// TIA Portal project "Mel7_new" (V15.1) (continued)
   L_1c_18."Индикатор: Обрыв" := FALSE;
   L_1c_18."Индикатор: В норме" := FALSE;
   L_1c_18."Индикатор: HH активирована" := FALSE;
   L_1c_18."Индикатор: H активирована" := FALSE;
   L_1c_18."Индикатор: L активирована" := FALSE;
   L_1c_18."Индикатор: LL активирована" := FALSE;
   L_1c_18."Уставка: MAX" := 450.0;
   L_1c_18."Уставка: MIN" := 0.0;
   L_1c_18."Уставка: HH" := 80.0;
   L_1c_18."Уставка: H" := 70.0;
   L_1c_18."Уставка: L" := 15.0;
   L_1c_18."Уставка: LL" := 10.0;
   L_1c_18."Уставка: Перелёт" := 20.0;
   L_1c_18."Уставка: Недолёт" := 4.0;
   L_1c_18.PV := 0.0813802;
   L_1c_18.Ток := 4.002893;
   L_1c_18.AnimCode := 0;
   L_1c_18.Error := 16#0000;
   L_1c_18.Bipolar := FALSE;
   L_1c_18.Overshoot_MIN := 27649;
   L_1c_18.Undershoot_MAX := -1;
   L_1c_19."Кнопка: Закрыть фейсплату" := FALSE;
   L_1c_19."Кнопка: Активировать HH" := FALSE;
   L_1c_19."Кнопка: Активировать H" := FALSE;
   L_1c_19."Кнопка: Активировать L" := FALSE;
   L_1c_19."Кнопка: Активировать LL" := FALSE;
   L_1c_19."Кнопка: Ремонт" := FALSE;
   L_1c_19.Видимость := FALSE;
   L_1c_19."Индикатор: Зашкал" := FALSE;
   L_1c_19."Индикатор: Перелёт" := FALSE;
   L_1c_19."Авария: Выход за HH" := FALSE;
   L_1c_19."Предупреждение: Выход за H" := FALSE;
   L_1c_19."Предупреждение: Выход за L" := FALSE;
   L_1c_19."Авария: Выход за LL" := FALSE;
   L_1c_19."Индикатор: Недолет" := FALSE;
   L_1c_19."Индикатор: Обрыв" := FALSE;
   L_1c_19."Индикатор: В норме" := FALSE;
   L_1c_19."Индикатор: HH активирована" := FALSE;
   L_1c_19."Индикатор: H активирована" := FALSE;
   L_1c_19."Индикатор: L активирована" := FALSE;
   L_1c_19."Индикатор: LL активирована" := FALSE;
   L_1c_19."Уставка: MAX" := 100.0;
   L_1c_19."Уставка: MIN" := 0.0;
   L_1c_19."Уставка: HH" := 80.0;
   L_1c_19."Уставка: H" := 70.0;
   L_1c_19."Уставка: L" := 15.0;
   L_1c_19."Уставка: LL" := 10.0;
   L_1c_19."Уставка: Перелёт" := 20.0;
   L_1c_19."Уставка: Недолёт" := 4.0;
   L_1c_19.PV := 0.1157407;
   L_1c_19.Ток := 4.018518;
   L_1c_19.AnimCode := 0;
   L_1c_19.Error := 16#0000;
   L_1c_19.Bipolar := FALSE;
   L_1c_19.Overshoot_MIN := 27649;
   L_1c_19.Undershoot_MAX := -1;
   L_1c_20."Кнопка: Закрыть фейсплату" := FALSE;
   L_1c_20."Кнопка: Активировать H" := FALSE;
   L_1c_20."Кнопка: Активировать L" := FALSE;
   L_1c_20."Кнопка: Активировать LL" := FALSE;
   L_1c_20."Кнопка: Ремонт" := FALSE;
   L_1c_20.Видимость := FALSE;
   L_1c_20."Индикатор: Зашкал" := FALSE;
   L_1c_20."Индикатор: Перелёт" := FALSE;
   L_1c_20."Авария: Выход за HH" := FALSE;
   L_1c_20."Предупреждение: Выход за H" := FALSE;
   L_1c_20."Предупреждение: Выход за L" := FALSE;
   L_1c_20."Авария: Выход за LL" := FALSE;
   L_1c_20."Индикатор: Недолет" := FALSE;
   L_1c_20."Индикатор: Обрыв" := FALSE;
   L_1c_20."Индикатор: В норме" := FALSE;
   L_1c_20."Индикатор: HH активирована" := FALSE;
   L_1c_20."Индикатор: H активирована" := FALSE;
   L_1c_20."Индикатор: L активирована" := FALSE;
   L_1c_20."Индикатор: LL активирована" := FALSE;
   L_1c_20."Уставка: MAX" := 100.0;
   L_1c_20."Уставка: MIN" := 0.0;
   L_1c_20."Уставка: HH" := 65.0;
   L_1c_20."Уставка: H" := 50.0;
   L_1c_20."Уставка: L" := 15.0;
   L_1c_20."Уставка: LL" := 10.0;
   L_1c_20."Уставка: Перелёт" := 20.0;
   L_1c_20."Уставка: Недолёт" := 4.0;
   L_1c_20.PV := 21.4;
   L_1c_20.Ток := 0.0;
   L_1c_20.AnimCode := 0;
   L_1c_20.Error := 16#0000;
   L_1c_20.Bipolar := FALSE;
   L_1c_20.Overshoot_MIN := 27649;
   L_1c_20.Undershoot_MAX := -1;
   L_1c_21."Кнопка: Закрыть фейсплату" := FALSE;
   L_1c_21."Кнопка: Активировать HH" := FALSE;
   L_1c_21."Кнопка: Активировать H" := FALSE;
   L_1c_21."Кнопка: Активировать L" := FALSE;
   L_1c_21."Кнопка: Активировать LL" := FALSE;
   L_1c_21."Кнопка: Ремонт" := FALSE;
   L_1c_21.Видимость := FALSE;
   L_1c_21."Индикатор: Зашкал" := FALSE;
   L_1c_21."Индикатор: Перелёт" := FALSE;
   L_1c_21."Авария: Выход за HH" := FALSE;
   L_1c_21."Предупреждение: Выход за H" := FALSE;
   L_1c_21."Предупреждение: Выход за L" := FALSE;
   L_1c_21."Авария: Выход за LL" := FALSE;
   L_1c_21."Индикатор: Недолет" := FALSE;
   L_1c_21."Индикатор: Обрыв" := FALSE;
   L_1c_21."Индикатор: В норме" := FALSE;
   L_1c_21."Индикатор: HH активирована" := FALSE;
   L_1c_21."Индикатор: H активирована" := FALSE;
   L_1c_21."Индикатор: L активирована" := FALSE;
   L_1c_21."Индикатор: LL активирована" := FALSE;
   L_1c_21."Уставка: MAX" := 100.0;
   L_1c_21."Уставка: MIN" := 0.0;
   L_1c_21."Уставка: HH" := 65.0;
   L_1c_21."Уставка: H" := 55.0;
   L_1c_21."Уставка: L" := 15.0;
   L_1c_21."Уставка: LL" := 10.0;
   L_1c_21."Уставка: Перелёт" := 20.0;
   L_1c_21."Уставка: Недолёт" := 4.0;
   L_1c_21.PV := 35.5;
   L_1c_21.Ток := 0.0;
   L_1c_21.AnimCode := 0;
   L_1c_21.Error := 16#0000;
   L_1c_21.Bipolar := FALSE;
   L_1c_21.Overshoot_MIN := 27649;
   L_1c_21.Undershoot_MAX := -1;
   L_1c_22."Кнопка: Закрыть фейсплату" := FALSE;
   L_1c_22."Кнопка: Активировать HH" := FALSE;
   L_1c_22."Кнопка: Активировать H" := FALSE;
   L_1c_22."Кнопка: Активировать L" := FALSE;
   L_1c_22."Кнопка: Активировать LL" := FALSE;
   L_1c_22."Кнопка: Ремонт" := FALSE;
   L_1c_22.Видимость := FALSE;
   L_1c_22."Индикатор: Зашкал" := FALSE;
   L_1c_22."Индикатор: Перелёт" := FALSE;
   L_1c_22."Авария: Выход за HH" := FALSE;
   L_1c_22."Предупреждение: Выход за H" := FALSE;
   L_1c_22."Предупреждение: Выход за L" := FALSE;
   L_1c_22."Авария: Выход за LL" := FALSE;
   L_1c_22."Индикатор: Недолет" := FALSE;
   L_1c_22."Индикатор: Обрыв" := FALSE;
   L_1c_22."Индикатор: В норме" := FALSE;
   L_1c_22."Индикатор: HH активирована" := FALSE;
   L_1c_22."Индикатор: H активирована" := FALSE;
   L_1c_22."Индикатор: L активирована" := FALSE;
   L_1c_22."Индикатор: LL активирована" := FALSE;
   L_1c_22."Уставка: MAX" := 100.0;
   L_1c_22."Уставка: MIN" := 0.0;
   L_1c_22."Уставка: HH" := 65.0;
   L_1c_22."Уставка: H" := 55.0;
   L_1c_22."Уставка: L" := 15.0;
   L_1c_22."Уставка: LL" := 10.0;
   L_1c_22."Уставка: Перелёт" := 20.0;
   L_1c_22."Уставка: Недолёт" := 4.0;
   L_1c_22.PV := 36.0;
   L_1c_22.Ток := 0.0;
   L_1c_22.AnimCode := 0;
   L_1c_22.Error := 16#0000;
   L_1c_22.Bipolar := FALSE;
   L_1c_22.Overshoot_MIN := 27649;
   L_1c_22.Undershoot_MAX := -1;
   L_1c_23."Кнопка: Закрыть фейсплату" := FALSE;
   L_1c_23."Кнопка: Активировать HH" := FALSE;
   L_1c_23."Кнопка: Активировать H" := FALSE;
   L_1c_23."Кнопка: Активировать L" := FALSE;
   L_1c_23."Кнопка: Активировать LL" := FALSE;
   L_1c_23."Кнопка: Ремонт" := FALSE;
   L_1c_23.Видимость := FALSE;
   L_1c_23."Индикатор: Зашкал" := FALSE;
   L_1c_23."Индикатор: Перелёт" := FALSE;
   L_1c_23."Авария: Выход за HH" := FALSE;
   L_1c_23."Предупреждение: Выход за H" := FALSE;
   L_1c_23."Предупреждение: Выход за L" := FALSE;
   L_1c_23."Авария: Выход за LL" := FALSE;
   L_1c_23."Индикатор: Недолет" := FALSE;
   L_1c_23."Индикатор: Обрыв" := FALSE;
   L_1c_23."Индикатор: В норме" := FALSE;
   L_1c_23."Индикатор: HH активирована" := FALSE;
   L_1c_23."Индикатор: H активирована" := FALSE;
   L_1c_23."Индикатор: L активирована" := FALSE;
   L_1c_23."Индикатор: LL активирована" := FALSE;
   L_1c_23."Уставка: MAX" := 100.0;
   L_1c_23."Уставка: MIN" := 0.0;
   L_1c_23."Уставка: HH" := 65.0;
   L_1c_23."Уставка: H" := 55.0;
   L_1c_23."Уставка: L" := 15.0;
   L_1c_23."Уставка: LL" := 10.0;
   L_1c_23."Уставка: Перелёт" := 20.0;
   L_1c_23."Уставка: Недолёт" := 4.0;
   L_1c_23.PV := 24.0;
   L_1c_23.Ток := 0.0;
   L_1c_23.AnimCode := 0;
   L_1c_23.Error := 16#0000;
   L_1c_23.Bipolar := FALSE;
   L_1c_23.Overshoot_MIN := 27649;
   L_1c_23.Undershoot_MAX := -1;
   L_1c_24."Кнопка: Закрыть фейсплату" := FALSE;
   L_1c_24."Кнопка: Активировать HH" := FALSE;
   L_1c_24."Кнопка: Активировать H" := FALSE;
   L_1c_24."Кнопка: Активировать L" := FALSE;
   L_1c_24."Кнопка: Активировать LL" := FALSE;
   L_1c_24."Кнопка: Ремонт" := FALSE;
   L_1c_24.Видимость := FALSE;
   L_1c_24."Индикатор: Зашкал" := FALSE;
   L_1c_24."Индикатор: Перелёт" := FALSE;
   L_1c_24."Авария: Выход за HH" := FALSE;
   L_1c_24."Предупреждение: Выход за H" := FALSE;
   L_1c_24."Предупреждение: Выход за L" := FALSE;
   L_1c_24."Авария: Выход за LL" := FALSE;
   L_1c_24."Индикатор: Недолет" := FALSE;
   L_1c_24."Индикатор: Обрыв" := FALSE;
   L_1c_24."Индикатор: В норме" := FALSE;
   L_1c_24."Индикатор: HH активирована" := FALSE;
   L_1c_24."Индикатор: H активирована" := FALSE;
   L_1c_24."Индикатор: L активирована" := FALSE;
   L_1c_24."Индикатор: LL активирована" := FALSE;
   L_1c_24."Уставка: MAX" := 100.0;
   L_1c_24."Уставка: MIN" := 0.0;
   L_1c_24."Уставка: HH" := 75.0;
   L_1c_24."Уставка: H" := 60.0;
   L_1c_24."Уставка: L" := 15.0;
   L_1c_24."Уставка: LL" := 10.0;
   L_1c_24."Уставка: Перелёт" := 20.0;
   L_1c_24."Уставка: Недолёт" := 4.0;
   L_1c_24.PV := 28.4;
   L_1c_24.Ток := 0.0;
   L_1c_24.AnimCode := 0;
   L_1c_24.Error := 16#0000;
   L_1c_24.Bipolar := FALSE;
   L_1c_24.Overshoot_MIN := 27649;
   L_1c_24.Undershoot_MAX := -1;
   L_1c_25."Кнопка: Закрыть фейсплату" := FALSE;
   L_1c_25."Кнопка: Активировать HH" := FALSE;
   L_1c_25."Кнопка: Активировать H" := FALSE;
   L_1c_25."Кнопка: Активировать L" := FALSE;
   L_1c_25."Кнопка: Активировать LL" := FALSE;
   L_1c_25."Кнопка: Ремонт" := FALSE;
   L_1c_25.Видимость := FALSE;
   L_1c_25."Индикатор: Зашкал" := FALSE;
   L_1c_25."Индикатор: Перелёт" := FALSE;
   L_1c_25."Авария: Выход за HH" := FALSE;
   L_1c_25."Предупреждение: Выход за H" := FALSE;
   L_1c_25."Предупреждение: Выход за L" := FALSE;
   L_1c_25."Авария: Выход за LL" := FALSE;
   L_1c_25."Индикатор: Недолет" := FALSE;
   L_1c_25."Индикатор: Обрыв" := FALSE;
   L_1c_25."Индикатор: В норме" := FALSE;
   L_1c_25."Индикатор: HH активирована" := FALSE;
   L_1c_25."Индикатор: H активирована" := FALSE;
   L_1c_25."Индикатор: L активирована" := FALSE;
   L_1c_25."Индикатор: LL активирована" := FALSE;
   L_1c_25."Уставка: MAX" := 100.0;
   L_1c_25."Уставка: MIN" := 0.0;
   L_1c_25."Уставка: HH" := 60.0;
   L_1c_25."Уставка: H" := 50.0;
   L_1c_25."Уставка: L" := 13.0;
   L_1c_25."Уставка: LL" := 10.0;
   L_1c_25."Уставка: Перелёт" := 20.0;
   L_1c_25."Уставка: Недолёт" := 4.0;
   L_1c_25.PV := 17.3;
   L_1c_25.Ток := 0.0;
   L_1c_25.AnimCode := 0;
   L_1c_25.Error := 16#0000;
   L_1c_25.Bipolar := FALSE;
   L_1c_25.Overshoot_MIN := 27649;
   L_1c_25.Undershoot_MAX := -1;
   L_1c_26."Кнопка: Закрыть фейсплату" := FALSE;
   L_1c_26."Кнопка: Активировать H" := FALSE;
   L_1c_26."Кнопка: Активировать L" := FALSE;
   L_1c_26."Кнопка: Активировать LL" := FALSE;
   L_1c_26."Кнопка: Ремонт" := FALSE;
   L_1c_26.Видимость := FALSE;
   L_1c_26."Индикатор: Зашкал" := FALSE;
   L_1c_26."Индикатор: Перелёт" := FALSE;
   L_1c_26."Авария: Выход за HH" := FALSE;
   L_1c_26."Предупреждение: Выход за H" := FALSE;
   L_1c_26."Предупреждение: Выход за L" := FALSE;
   L_1c_26."Авария: Выход за LL" := FALSE;
   L_1c_26."Индикатор: Недолет" := FALSE;
   L_1c_26."Индикатор: Обрыв" := FALSE;
   L_1c_26."Индикатор: В норме" := FALSE;
   L_1c_26."Индикатор: HH активирована" := FALSE;
   L_1c_26."Индикатор: H активирована" := FALSE;
   L_1c_26."Индикатор: L активирована" := FALSE;
   L_1c_26."Индикатор: LL активирована" := FALSE;
   L_1c_26."Уставка: MAX" := 100.0;
   L_1c_26."Уставка: MIN" := 0.0;
   L_1c_26."Уставка: HH" := 60.0;
   L_1c_26."Уставка: H" := 50.0;
   L_1c_26."Уставка: L" := 15.0;
   L_1c_26."Уставка: LL" := 10.0;
   L_1c_26."Уставка: Перелёт" := 20.0;
   L_1c_26."Уставка: Недолёт" := 4.0;
   L_1c_26.PV := 18.5;
   L_1c_26.Ток := 0.0;
   L_1c_26.AnimCode := 0;
   L_1c_26.Error := 16#0000;
   L_1c_26.Bipolar := FALSE;
   L_1c_26.Overshoot_MIN := 27649;
   L_1c_26.Undershoot_MAX := -1;
   L_1c_27."Кнопка: Закрыть фейсплату" := FALSE;
   L_1c_27."Кнопка: Активировать HH" := FALSE;
   L_1c_27."Кнопка: Активировать H" := FALSE;
   L_1c_27."Кнопка: Активировать L" := FALSE;
   L_1c_27."Кнопка: Активировать LL" := FALSE;
   L_1c_27."Кнопка: Ремонт" := FALSE;
   L_1c_27.Видимость := FALSE;
   L_1c_27."Индикатор: Зашкал" := FALSE;
   L_1c_27."Индикатор: Перелёт" := FALSE;
   L_1c_27."Авария: Выход за HH" := FALSE;
   L_1c_27."Предупреждение: Выход за H" := FALSE;
   L_1c_27."Предупреждение: Выход за L" := FALSE;
   L_1c_27."Авария: Выход за LL" := FALSE;
   L_1c_27."Индикатор: Недолет" := FALSE;
   L_1c_27."Индикатор: Обрыв" := FALSE;
   L_1c_27."Индикатор: В норме" := FALSE;
   L_1c_27."Индикатор: HH активирована" := FALSE;
   L_1c_27."Индикатор: H активирована" := FALSE;
   L_1c_27."Индикатор: L активирована" := FALSE;
   L_1c_27."Индикатор: LL активирована" := FALSE;
   L_1c_27."Уставка: MAX" := 100.0;
   L_1c_27."Уставка: MIN" := 0.0;
   L_1c_27."Уставка: HH" := 60.0;
   L_1c_27."Уставка: H" := 50.0;
   L_1c_27."Уставка: L" := 15.0;
   L_1c_27."Уставка: LL" := 10.0;
   L_1c_27."Уставка: Перелёт" := 20.0;
   L_1c_27."Уставка: Недолёт" := 4.0;
   L_1c_27.PV := 18.6;
   L_1c_27.Ток := 0.0;
   L_1c_27.AnimCode := 0;
   L_1c_27.Error := 16#0000;
   L_1c_27.Bipolar := FALSE;
   L_1c_27.Overshoot_MIN := 27649;
   L_1c_27.Undershoot_MAX := -1;
   L_1c_28."Кнопка: Закрыть фейсплату" := FALSE;
   L_1c_28."Кнопка: Активировать HH" := FALSE;
   L_1c_28."Кнопка: Активировать H" := FALSE;
   L_1c_28."Кнопка: Активировать L" := FALSE;
   L_1c_28."Кнопка: Активировать LL" := FALSE;
   L_1c_28."Кнопка: Ремонт" := FALSE;
   L_1c_28.Видимость := FALSE;
   L_1c_28."Индикатор: Зашкал" := FALSE;
   L_1c_28."Индикатор: Перелёт" := FALSE;
   L_1c_28."Авария: Выход за HH" := FALSE;
   L_1c_28."Предупреждение: Выход за H" := FALSE;
   L_1c_28."Предупреждение: Выход за L" := FALSE;
   L_1c_28."Авария: Выход за LL" := FALSE;
   L_1c_28."Индикатор: Недолет" := FALSE;
   L_1c_28."Индикатор: Обрыв" := FALSE;
   L_1c_28."Индикатор: В норме" := FALSE;
   L_1c_28."Индикатор: HH активирована" := FALSE;
   L_1c_28."Индикатор: H активирована" := FALSE;
   L_1c_28."Индикатор: L активирована" := FALSE;
   L_1c_28."Индикатор: LL активирована" := FALSE;
   L_1c_28."Уставка: MAX" := 100.0;
   L_1c_28."Уставка: MIN" := 0.0;
   L_1c_28."Уставка: HH" := 80.0;
   L_1c_28."Уставка: H" := 70.0;
   L_1c_28."Уставка: L" := 15.0;
   L_1c_28."Уставка: LL" := 10.0;
   L_1c_28."Уставка: Перелёт" := 20.0;
   L_1c_28."Уставка: Недолёт" := 4.0;
   L_1c_28.PV := 0.01808449;
   L_1c_28.Ток := 4.002893;
   L_1c_28.AnimCode := 0;
   L_1c_28.Error := 16#0000;
   L_1c_28.Bipolar := FALSE;
   L_1c_28.Overshoot_MIN := 27649;
   L_1c_28.Undershoot_MAX := -1;
   L_1c_29."Кнопка: Закрыть фейсплату" := FALSE;
   L_1c_29."Кнопка: Активировать HH" := FALSE;
   L_1c_29."Кнопка: Активировать H" := FALSE;
   L_1c_29."Кнопка: Активировать L" := FALSE;
   L_1c_29."Кнопка: Активировать LL" := FALSE;
   L_1c_29."Кнопка: Ремонт" := FALSE;
   L_1c_29.Видимость := FALSE;
   L_1c_29."Индикатор: Зашкал" := FALSE;
   L_1c_29."Индикатор: Перелёт" := FALSE;
   L_1c_29."Авария: Выход за HH" := FALSE;
   L_1c_29."Предупреждение: Выход за H" := FALSE;
   L_1c_29."Предупреждение: Выход за L" := FALSE;
   L_1c_29."Авария: Выход за LL" := FALSE;
   L_1c_29."Индикатор: Недолет" := FALSE;
   L_1c_29."Индикатор: Обрыв" := FALSE;
   L_1c_29."Индикатор: В норме" := FALSE;
   L_1c_29."Индикатор: HH активирована" := FALSE;
   L_1c_29."Индикатор: H активирована" := FALSE;
   L_1c_29."Индикатор: L активирована" := FALSE;
   L_1c_29."Индикатор: LL активирована" := FALSE;
   L_1c_29."Уставка: MAX" := 100.0;
   L_1c_29."Уставка: MIN" := 0.0;
   L_1c_29."Уставка: HH" := 75.0;
   L_1c_29."Уставка: H" := 50.0;
   L_1c_29."Уставка: L" := 15.0;
   L_1c_29."Уставка: LL" := 10.0;
   L_1c_29."Уставка: Перелёт" := 20.0;
   L_1c_29."Уставка: Недолёт" := 4.0;
   L_1c_29.PV := 24.5;
   L_1c_29.Ток := 0.0;
   L_1c_29.AnimCode := 0;
   L_1c_29.Error := 16#0000;
   L_1c_29.Bipolar := FALSE;
   L_1c_29.Overshoot_MIN := 27649;
   L_1c_29.Undershoot_MAX := -1;
   L_1c_30."Кнопка: Закрыть фейсплату" := FALSE;
   L_1c_30."Кнопка: Активировать HH" := FALSE;
   L_1c_30."Кнопка: Активировать H" := FALSE;
   L_1c_30."Кнопка: Активировать L" := FALSE;
   L_1c_30."Кнопка: Активировать LL" := FALSE;
   L_1c_30."Кнопка: Ремонт" := FALSE;
   L_1c_30.Видимость := FALSE;
   L_1c_30."Индикатор: Зашкал" := FALSE;
   L_1c_30."Индикатор: Перелёт" := FALSE;
   L_1c_30."Авария: Выход за HH" := FALSE;
   L_1c_30."Предупреждение: Выход за H" := FALSE;
   L_1c_30."Предупреждение: Выход за L" := FALSE;
   L_1c_30."Авария: Выход за LL" := FALSE;
   L_1c_30."Индикатор: Недолет" := FALSE;
   L_1c_30."Индикатор: Обрыв" := FALSE;
   L_1c_30."Индикатор: В норме" := FALSE;
   L_1c_30."Индикатор: HH активирована" := FALSE;
   L_1c_30."Индикатор: H активирована" := FALSE;
   L_1c_30."Индикатор: L активирована" := FALSE;
   L_1c_30."Индикатор: LL активирована" := FALSE;
   L_1c_30."Уставка: MAX" := 100.0;
   L_1c_30."Уставка: MIN" := 0.0;
   L_1c_30."Уставка: HH" := 80.0;
   L_1c_30."Уставка: H" := 70.0;
   L_1c_30."Уставка: L" := 15.0;
   L_1c_30."Уставка: LL" := 10.0;
   L_1c_30."Уставка: Перелёт" := 20.0;
   L_1c_30."Уставка: Недолёт" := 4.0;
   L_1c_30.PV := 0.1482928;
   L_1c_30.Ток := 4.023727;
   L_1c_30.AnimCode := 0;
   L_1c_30.Error := 16#0000;
   L_1c_30.Bipolar := FALSE;
   L_1c_30.Overshoot_MIN := 27649;
   L_1c_30.Undershoot_MAX := -1;
   L_1c_31."Кнопка: Закрыть фейсплату" := FALSE;
   L_1c_31."Кнопка: Активировать HH" := FALSE;
   L_1c_31."Кнопка: Активировать H" := FALSE;
   L_1c_31."Кнопка: Активировать L" := FALSE;
   L_1c_31."Кнопка: Активировать LL" := FALSE;
   L_1c_31."Кнопка: Ремонт" := FALSE;
   L_1c_31.Видимость := FALSE;
   L_1c_31."Индикатор: Зашкал" := FALSE;
   L_1c_31."Индикатор: Перелёт" := FALSE;
   L_1c_31."Авария: Выход за HH" := FALSE;
   L_1c_31."Предупреждение: Выход за H" := FALSE;
   L_1c_31."Предупреждение: Выход за L" := FALSE;
   L_1c_31."Авария: Выход за LL" := FALSE;
   L_1c_31."Индикатор: Недолет" := FALSE;
   L_1c_31."Индикатор: Обрыв" := FALSE;
   L_1c_31."Индикатор: В норме" := FALSE;
   L_1c_31."Индикатор: HH активирована" := FALSE;
   L_1c_31."Индикатор: H активирована" := FALSE;
   L_1c_31."Индикатор: L активирована" := FALSE;
   L_1c_31."Индикатор: LL активирована" := FALSE;
   L_1c_31."Уставка: MAX" := 100.0;
   L_1c_31."Уставка: MIN" := 0.0;
   L_1c_31."Уставка: HH" := 80.0;
   L_1c_31."Уставка: H" := 70.0;
   L_1c_31."Уставка: L" := 15.0;
   L_1c_31."Уставка: LL" := 10.0;
   L_1c_31."Уставка: Перелёт" := 20.0;
   L_1c_31."Уставка: Недолёт" := 4.0;
   L_1c_31.PV := 0.07595486;
   L_1c_31.Ток := 4.012153;
   L_1c_31.AnimCode := 0;
   L_1c_31.Error := 16#0000;
   L_1c_31.Bipolar := FALSE;
   L_1c_31.Overshoot_MIN := 27649;
   L_1c_31.Undershoot_MAX := -1;
   L_1c_32."Кнопка: Закрыть фейсплату" := FALSE;
   L_1c_32."Кнопка: Активировать HH" := FALSE;
   L_1c_32."Кнопка: Активировать H" := FALSE;
   L_1c_32."Кнопка: Активировать L" := FALSE;
   L_1c_32."Кнопка: Активировать LL" := FALSE;
   L_1c_32."Кнопка: Ремонт" := FALSE;
   L_1c_32.Видимость := FALSE;
   L_1c_32."Индикатор: Зашкал" := FALSE;
   L_1c_32."Индикатор: Перелёт" := FALSE;
   L_1c_32."Авария: Выход за HH" := FALSE;
   L_1c_32."Предупреждение: Выход за H" := FALSE;
   L_1c_32."Предупреждение: Выход за L" := FALSE;
   L_1c_32."Авария: Выход за LL" := FALSE;
   L_1c_32."Индикатор: Недолет" := FALSE;
   L_1c_32."Индикатор: Обрыв" := FALSE;
   L_1c_32."Индикатор: В норме" := FALSE;
   L_1c_32."Индикатор: HH активирована" := FALSE;
   L_1c_32."Индикатор: H активирована" := FALSE;
   L_1c_32."Индикатор: L активирована" := FALSE;
   L_1c_32."Индикатор: LL активирована" := FALSE;
   L_1c_32."Уставка: MAX" := 1000.0;
   L_1c_32."Уставка: MIN" := 0.0;
   L_1c_32."Уставка: HH" := 80.0;
   L_1c_32."Уставка: H" := 70.0;
   L_1c_32."Уставка: L" := 15.0;
   L_1c_32."Уставка: LL" := 10.0;
   L_1c_32."Уставка: Перелёт" := 20.0;
   L_1c_32."Уставка: Недолёт" := 4.0;
   L_1c_32.PV := 40.76244;
   L_1c_32.Ток := 4.652199;
   L_1c_32.AnimCode := 0;
   L_1c_32.Error := 16#0000;
   L_1c_32.Bipolar := FALSE;
   L_1c_32.Overshoot_MIN := 27649;
   L_1c_32.Undershoot_MAX := -1;
   L_1c_33."Кнопка: Закрыть фейсплату" := FALSE;
   L_1c_33."Кнопка: Активировать HH" := FALSE;
   L_1c_33."Кнопка: Активировать H" := FALSE;
   L_1c_33."Кнопка: Активировать L" := FALSE;
   L_1c_33."Кнопка: Активировать LL" := FALSE;
   L_1c_33."Кнопка: Ремонт" := FALSE;
   L_1c_33.Видимость := FALSE;
   L_1c_33."Индикатор: Зашкал" := FALSE;
   L_1c_33."Индикатор: Перелёт" := FALSE;
   L_1c_33."Авария: Выход за HH" := FALSE;
   L_1c_33."Предупреждение: Выход за H" := FALSE;
   L_1c_33."Предупреждение: Выход за L" := FALSE;
   L_1c_33."Авария: Выход за LL" := FALSE;
   L_1c_33."Индикатор: Недолет" := FALSE;
   L_1c_33."Индикатор: Обрыв" := FALSE;
   L_1c_33."Индикатор: В норме" := FALSE;
   L_1c_33."Индикатор: HH активирована" := FALSE;
   L_1c_33."Индикатор: H активирована" := FALSE;
   L_1c_33."Индикатор: L активирована" := FALSE;
   L_1c_33."Индикатор: LL активирована" := FALSE;
   L_1c_33."Уставка: MAX" := 1000.0;
   L_1c_33."Уставка: MIN" := 0.0;
   L_1c_33."Уставка: HH" := 80.0;
   L_1c_33."Уставка: H" := 70.0;
   L_1c_33."Уставка: L" := 15.0;
   L_1c_33."Уставка: LL" := 10.0;
   L_1c_33."Уставка: Перелёт" := 20.0;
   L_1c_33."Уставка: Недолёт" := 4.0;
   L_1c_33.PV := 35.66262;
   L_1c_33.Ток := 4.570602;
   L_1c_33.AnimCode := 0;
   L_1c_33.Error := 16#0000;
   L_1c_33.Bipolar := FALSE;
   L_1c_33.Overshoot_MIN := 27649;
   L_1c_33.Undershoot_MAX := -1;
   L_1c_36."Кнопка: Закрыть фейсплату" := FALSE;
   L_1c_36."Кнопка: Активировать HH" := FALSE;
   L_1c_36."Кнопка: Активировать H" := FALSE;
   L_1c_36."Кнопка: Активировать L" := FALSE;
   L_1c_36."Кнопка: Активировать LL" := FALSE;
   L_1c_36."Кнопка: Ремонт" := FALSE;
   L_1c_36.Видимость := FALSE;
   L_1c_36."Индикатор: Зашкал" := FALSE;
   L_1c_36."Индикатор: Перелёт" := FALSE;
   L_1c_36."Авария: Выход за HH" := FALSE;
   L_1c_36."Предупреждение: Выход за H" := FALSE;
   L_1c_36."Предупреждение: Выход за L" := FALSE;
   L_1c_36."Авария: Выход за LL" := FALSE;
   L_1c_36."Индикатор: Недолет" := TRUE;
   L_1c_36."Индикатор: Обрыв" := FALSE;
   L_1c_36."Индикатор: В норме" := FALSE;
   L_1c_36."Индикатор: HH активирована" := FALSE;
   L_1c_36."Индикатор: H активирована" := FALSE;
   L_1c_36."Индикатор: L активирована" := FALSE;
   L_1c_36."Индикатор: LL активирована" := FALSE;
   L_1c_36."Уставка: MAX" := 50.0;
   L_1c_36."Уставка: MIN" := 0.0;
   L_1c_36."Уставка: HH" := 80.0;
   L_1c_36."Уставка: H" := 70.0;
   L_1c_36."Уставка: L" := 15.0;
   L_1c_36."Уставка: LL" := 10.0;
   L_1c_36."Уставка: Перелёт" := 20.0;
   L_1c_36."Уставка: Недолёт" := 4.0;
   L_1c_36.PV := -1.114005;
   L_1c_36.Ток := 3.643518;
   L_1c_36.AnimCode := 2;
   L_1c_36.Error := 16#0000;
   L_1c_36.Bipolar := FALSE;
   L_1c_36.Overshoot_MIN := 27649;
   L_1c_36.Undershoot_MAX := -1;
   L_1c_37."Кнопка: Закрыть фейсплату" := FALSE;
   L_1c_37."Кнопка: Активировать HH" := FALSE;
   L_1c_37."Кнопка: Активировать H" := FALSE;
   L_1c_37."Кнопка: Активировать L" := FALSE;
   L_1c_37."Кнопка: Активировать LL" := FALSE;
   L_1c_37."Кнопка: Ремонт" := FALSE;
   L_1c_37.Видимость := FALSE;
   L_1c_37."Индикатор: Зашкал" := FALSE;
   L_1c_37."Индикатор: Перелёт" := FALSE;
   L_1c_37."Авария: Выход за HH" := FALSE;
   L_1c_37."Предупреждение: Выход за H" := FALSE;
   L_1c_37."Предупреждение: Выход за L" := FALSE;
   L_1c_37."Авария: Выход за LL" := FALSE;
   L_1c_37."Индикатор: Недолет" := TRUE;
   L_1c_37."Индикатор: Обрыв" := FALSE;
   L_1c_37."Индикатор: В норме" := FALSE;
   L_1c_37."Индикатор: HH активирована" := FALSE;
   L_1c_37."Индикатор: H активирована" := FALSE;
   L_1c_37."Индикатор: L активирована" := FALSE;
   L_1c_37."Индикатор: LL активирована" := FALSE;
   L_1c_37."Уставка: MAX" := 100.0;
   L_1c_37."Уставка: MIN" := 0.0;
   L_1c_37."Уставка: HH" := 80.0;
   L_1c_37."Уставка: H" := 70.0;
   L_1c_37."Уставка: L" := 15.0;
   L_1c_37."Уставка: LL" := 10.0;
   L_1c_37."Уставка: Перелёт" := 20.0;
   L_1c_37."Уставка: Недолёт" := 4.0;
   L_1c_37.PV := -0.2531829;
   L_1c_37.Ток := 3.959491;
   L_1c_37.AnimCode := 2;
   L_1c_37.Error := 16#0000;
   L_1c_37.Bipolar := FALSE;
   L_1c_37.Overshoot_MIN := 27649;
   L_1c_37.Undershoot_MAX := -1;
   L_1c_38."Кнопка: Закрыть фейсплату" := FALSE;
   L_1c_38."Кнопка: Активировать HH" := FALSE;
   L_1c_38."Кнопка: Активировать H" := FALSE;
   L_1c_38."Кнопка: Активировать L" := FALSE;
   L_1c_38."Кнопка: Активировать LL" := FALSE;
   L_1c_38."Кнопка: Ремонт" := FALSE;
   L_1c_38.Видимость := FALSE;
   L_1c_38."Индикатор: Зашкал" := FALSE;
   L_1c_38."Индикатор: Перелёт" := FALSE;
   L_1c_38."Авария: Выход за HH" := FALSE;
   L_1c_38."Предупреждение: Выход за H" := FALSE;
   L_1c_38."Предупреждение: Выход за L" := FALSE;
   L_1c_38."Авария: Выход за LL" := FALSE;
   L_1c_38."Индикатор: Недолет" := TRUE;
   L_1c_38."Индикатор: Обрыв" := FALSE;
   L_1c_38."Индикатор: В норме" := FALSE;
   L_1c_38."Индикатор: HH активирована" := FALSE;
   L_1c_38."Индикатор: H активирована" := FALSE;
   L_1c_38."Индикатор: L активирована" := FALSE;
   L_1c_38."Индикатор: LL активирована" := FALSE;
   L_1c_38."Уставка: MAX" := 100.0;
   L_1c_38."Уставка: MIN" := 0.0;
   L_1c_38."Уставка: HH" := 80.0;
   L_1c_38."Уставка: H" := 70.0;
   L_1c_38."Уставка: L" := 15.0;
   L_1c_38."Уставка: LL" := 10.0;
   L_1c_38."Уставка: Перелёт" := 20.0;
   L_1c_38."Уставка: Недолёт" := 4.0;
   L_1c_38.PV := -0.7559317;
   L_1c_38.Ток := 3.879051;
   L_1c_38.AnimCode := 2;
   L_1c_38.Error := 16#0000;
   L_1c_38.Bipolar := FALSE;
   L_1c_38.Overshoot_MIN := 27649;
   L_1c_38.Undershoot_MAX := -1;
   L_1c_39."Кнопка: Закрыть фейсплату" := FALSE;
   L_1c_39."Кнопка: Активировать HH" := FALSE;
   L_1c_39."Кнопка: Активировать H" := FALSE;
   L_1c_39."Кнопка: Активировать L" := FALSE;
   L_1c_39."Кнопка: Активировать LL" := FALSE;
   L_1c_39."Кнопка: Ремонт" := FALSE;
   L_1c_39.Видимость := FALSE;
   L_1c_39."Индикатор: Зашкал" := FALSE;
   L_1c_39."Индикатор: Перелёт" := FALSE;
   L_1c_39."Авария: Выход за HH" := FALSE;
   L_1c_39."Предупреждение: Выход за H" := FALSE;
   L_1c_39."Предупреждение: Выход за L" := FALSE;
   L_1c_39."Авария: Выход за LL" := FALSE;
   L_1c_39."Индикатор: Недолет" := FALSE;
   L_1c_39."Индикатор: Обрыв" := FALSE;
   L_1c_39."Индикатор: В норме" := FALSE;
   L_1c_39."Индикатор: HH активирована" := FALSE;
   L_1c_39."Индикатор: H активирована" := FALSE;
   L_1c_39."Индикатор: L активирована" := FALSE;
   L_1c_39."Индикатор: LL активирована" := FALSE;
   L_1c_39."Уставка: MAX" := 100.0;
   L_1c_39."Уставка: MIN" := 0.0;
   L_1c_39."Уставка: HH" := 80.0;
   L_1c_39."Уставка: H" := 70.0;
   L_1c_39."Уставка: L" := 15.0;
   L_1c_39."Уставка: LL" := 10.0;
   L_1c_39."Уставка: Перелёт" := 20.0;
   L_1c_39."Уставка: Недолёт" := 4.0;
   L_1c_39.PV := 0.0;
   L_1c_39.Ток := 4.0;
   L_1c_39.AnimCode := 0;
   L_1c_39.Error := 16#0000;
   L_1c_39.Bipolar := FALSE;
   L_1c_39.Overshoot_MIN := 27649;
   L_1c_39.Undershoot_MAX := -1;
   L_1c_40."Кнопка: Закрыть фейсплату" := FALSE;
   L_1c_40."Кнопка: Активировать HH" := FALSE;
   L_1c_40."Кнопка: Активировать H" := FALSE;
   L_1c_40."Кнопка: Активировать L" := FALSE;
   L_1c_40."Кнопка: Активировать LL" := FALSE;
   L_1c_40."Кнопка: Ремонт" := FALSE;
   L_1c_40.Видимость := FALSE;
   L_1c_40."Индикатор: Зашкал" := FALSE;
   L_1c_40."Индикатор: Перелёт" := FALSE;
   L_1c_40."Авария: Выход за HH" := FALSE;
   L_1c_40."Предупреждение: Выход за H" := FALSE;
   L_1c_40."Предупреждение: Выход за L" := FALSE;
   L_1c_40."Авария: Выход за LL" := FALSE;
   L_1c_40."Индикатор: Недолет" := FALSE;
   L_1c_40."Индикатор: Обрыв" := FALSE;
   L_1c_40."Индикатор: В норме" := FALSE;
   L_1c_40."Индикатор: HH активирована" := FALSE;
   L_1c_40."Индикатор: H активирована" := FALSE;
   L_1c_40."Индикатор: L активирована" := FALSE;
   L_1c_40."Индикатор: LL активирована" := FALSE;
   L_1c_40."Уставка: MAX" := 100.0;
   L_1c_40."Уставка: MIN" := 0.0;
   L_1c_40."Уставка: HH" := 80.0;
   L_1c_40."Уставка: H" := 70.0;
   L_1c_40."Уставка: L" := 15.0;
   L_1c_40."Уставка: LL" := 10.0;
   L_1c_40."Уставка: Перелёт" := 20.0;
   L_1c_40."Уставка: Недолёт" := 4.0;
   L_1c_40.PV := 0.4376447;
   L_1c_40.Ток := 4.070023;
   L_1c_40.AnimCode := 0;
   L_1c_40.Error := 16#0000;
   L_1c_40.Bipolar := FALSE;
   L_1c_40.Overshoot_MIN := 27649;
   L_1c_40.Undershoot_MAX := -1;
   L_1c_41."Кнопка: Закрыть фейсплату" := FALSE;
   L_1c_41."Кнопка: Активировать HH" := FALSE;
   L_1c_41."Кнопка: Активировать H" := FALSE;
   L_1c_41."Кнопка: Активировать L" := FALSE;
   L_1c_41."Кнопка: Активировать LL" := FALSE;
   L_1c_41."Кнопка: Ремонт" := FALSE;
   L_1c_41.Видимость := FALSE;
   L_1c_41."Индикатор: Зашкал" := FALSE;
   L_1c_41."Индикатор: Перелёт" := FALSE;
   L_1c_41."Авария: Выход за HH" := FALSE;
   L_1c_41."Предупреждение: Выход за H" := FALSE;
   L_1c_41."Предупреждение: Выход за L" := FALSE;
   L_1c_41."Авария: Выход за LL" := FALSE;
   L_1c_41."Индикатор: Недолет" := FALSE;
   L_1c_41."Индикатор: Обрыв" := FALSE;
   L_1c_41."Индикатор: В норме" := FALSE;
   L_1c_41."Индикатор: HH активирована" := FALSE;
   L_1c_41."Индикатор: H активирована" := FALSE;
   L_1c_41."Индикатор: L активирована" := FALSE;
   L_1c_41."Индикатор: LL активирована" := FALSE;
   L_1c_41."Уставка: MAX" := 100.0;
   L_1c_41."Уставка: MIN" := 0.0;
   L_1c_41."Уставка: HH" := 80.0;
   L_1c_41."Уставка: H" := 70.0;
   L_1c_41."Уставка: L" := 15.0;
   L_1c_41."Уставка: LL" := 10.0;
   L_1c_41."Уставка: Перелёт" := 20.0;
   L_1c_41."Уставка: Недолёт" := 4.0;
   L_1c_41.PV := 0.05063657;
   L_1c_41.Ток := 4.008102;
   L_1c_41.AnimCode := 0;
   L_1c_41.Error := 16#0000;
   L_1c_41.Bipolar := FALSE;
   L_1c_41.Overshoot_MIN := 27649;
   L_1c_41.Undershoot_MAX := -1;
   L_1c_42."Кнопка: Закрыть фейсплату" := FALSE;
   L_1c_42."Кнопка: Активировать HH" := FALSE;
   L_1c_42."Кнопка: Активировать H" := FALSE;
   L_1c_42."Кнопка: Активировать L" := FALSE;
   L_1c_42."Кнопка: Активировать LL" := FALSE;
   L_1c_42."Кнопка: Ремонт" := FALSE;
   L_1c_42.Видимость := FALSE;
   L_1c_42."Индикатор: Зашкал" := FALSE;
   L_1c_42."Индикатор: Перелёт" := FALSE;
   L_1c_42."Авария: Выход за HH" := FALSE;
   L_1c_42."Предупреждение: Выход за H" := FALSE;
   L_1c_42."Предупреждение: Выход за L" := FALSE;
   L_1c_42."Авария: Выход за LL" := FALSE;
   L_1c_42."Индикатор: Недолет" := FALSE;
   L_1c_42."Индикатор: Обрыв" := FALSE;
   L_1c_42."Индикатор: В норме" := FALSE;
   L_1c_42."Индикатор: HH активирована" := FALSE;
   L_1c_42."Индикатор: H активирована" := FALSE;
   L_1c_42."Индикатор: L активирована" := FALSE;
   L_1c_42."Индикатор: LL активирована" := FALSE;
   L_1c_42."Уставка: MAX" := 100.0;
   L_1c_42."Уставка: MIN" := 0.0;
   L_1c_42."Уставка: HH" := 80.0;
   L_1c_42."Уставка: H" := 70.0;
   L_1c_42."Уставка: L" := 15.0;
   L_1c_42."Уставка: LL" := 10.0;
   L_1c_42."Уставка: Перелёт" := 20.0;
   L_1c_42."Уставка: Недолёт" := 4.0;
   L_1c_42.PV := 0.06872106;
   L_1c_42.Ток := 4.010995;
   L_1c_42.AnimCode := 0;
   L_1c_42.Error := 16#0000;
   L_1c_42.Bipolar := FALSE;
   L_1c_42.Overshoot_MIN := 27649;
   L_1c_42.Undershoot_MAX := -1;
   L_1c_43."Уставка: MAX" := 65.0;
   L_1c_44."Уставка: MAX" := 65.0;
   L_1c_43."Кнопка: Закрыть фейсплату" := FALSE;
   L_1c_43."Кнопка: Активировать HH" := FALSE;
   L_1c_43."Кнопка: Активировать H" := FALSE;
   L_1c_43."Кнопка: Активировать L" := FALSE;
   L_1c_43."Кнопка: Активировать LL" := FALSE;
   L_1c_43."Кнопка: Ремонт" := FALSE;
   L_1c_43.Видимость := FALSE;
   L_1c_43."Индикатор: Зашкал" := FALSE;
   L_1c_43."Индикатор: Перелёт" := FALSE;
   L_1c_43."Авария: Выход за HH" := FALSE;
   L_1c_43."Предупреждение: Выход за H" := FALSE;
   L_1c_43."Предупреждение: Выход за L" := FALSE;
   L_1c_43."Авария: Выход за LL" := FALSE;
   L_1c_43."Индикатор: Недолет" := FALSE;
   L_1c_43."Индикатор: Обрыв" := FALSE;
   L_1c_43."Индикатор: В норме" := FALSE;
   L_1c_43."Индикатор: HH активирована" := FALSE;
   L_1c_43."Индикатор: H активирована" := FALSE;
   L_1c_43."Индикатор: L активирована" := FALSE;
   L_1c_43."Индикатор: LL активирована" := FALSE;
   L_1c_43."Уставка: MIN" := 0.0;
   L_1c_43."Уставка: HH" := 80.0;
   L_1c_43."Уставка: H" := 70.0;
   L_1c_43."Уставка: L" := 5.0;
   L_1c_43."Уставка: LL" := 10.0;
   L_1c_43."Уставка: Перелёт" := 20.0;
   L_1c_43."Уставка: Недолёт" := 4.0;
   L_1c_43.PV := 0.0;
   L_1c_43.Ток := 4.0;
   L_1c_43.AnimCode := 0;
   L_1c_43.Error := 16#0000;
   L_1c_43.Bipolar := FALSE;
   L_1c_43.Overshoot_MIN := 27649;
   L_1c_43.Undershoot_MAX := -1;
   L_1c_44."Кнопка: Закрыть фейсплату" := FALSE;
   L_1c_44."Кнопка: Активировать HH" := FALSE;
   L_1c_44."Кнопка: Активировать H" := FALSE;
   L_1c_44."Кнопка: Активировать L" := FALSE;
   L_1c_44."Кнопка: Активировать LL" := FALSE;
   L_1c_44."Кнопка: Ремонт" := FALSE;
   L_1c_44.Видимость := FALSE;
   L_1c_44."Индикатор: Зашкал" := FALSE;
   L_1c_44."Индикатор: Перелёт" := FALSE;
   L_1c_44."Авария: Выход за HH" := FALSE;
   L_1c_44."Предупреждение: Выход за H" := FALSE;
   L_1c_44."Предупреждение: Выход за L" := FALSE;
   L_1c_44."Авария: Выход за LL" := FALSE;
   L_1c_44."Индикатор: Недолет" := TRUE;
   L_1c_44."Индикатор: Обрыв" := FALSE;
   L_1c_44."Индикатор: В норме" := FALSE;
   L_1c_44."Индикатор: HH активирована" := FALSE;
   L_1c_44."Индикатор: H активирована" := FALSE;
   L_1c_44."Индикатор: L активирована" := FALSE;
   L_1c_44."Индикатор: LL активирована" := FALSE;
   L_1c_44."Уставка: MIN" := 0.0;
   L_1c_44."Уставка: HH" := 80.0;
   L_1c_44."Уставка: H" := 70.0;
   L_1c_44."Уставка: L" := 15.0;
   L_1c_44."Уставка: LL" := 10.0;
   L_1c_44."Уставка: Перелёт" := 20.0;
   L_1c_44."Уставка: Недолёт" := 4.0;
   L_1c_44.PV := -0.004701968;
   L_1c_44.Ток := 3.998842;
   L_1c_44.AnimCode := 2;
   L_1c_44.Error := 16#0000;
   L_1c_44.Bipolar := FALSE;
   L_1c_44.Overshoot_MIN := 27649;
   L_1c_44.Undershoot_MAX := -1;
   L_1c_45."Кнопка: Закрыть фейсплату" := FALSE;
   L_1c_45."Кнопка: Активировать HH" := FALSE;
   L_1c_45."Кнопка: Активировать H" := FALSE;
   L_1c_45."Кнопка: Активировать L" := FALSE;
   L_1c_45."Кнопка: Активировать LL" := FALSE;
   L_1c_45."Кнопка: Ремонт" := FALSE;
   L_1c_45.Видимость := FALSE;
   L_1c_45."Индикатор: Зашкал" := FALSE;
   L_1c_45."Индикатор: Перелёт" := FALSE;
   L_1c_45."Авария: Выход за HH" := FALSE;
   L_1c_45."Предупреждение: Выход за H" := FALSE;
   L_1c_45."Предупреждение: Выход за L" := FALSE;
   L_1c_45."Авария: Выход за LL" := FALSE;
   L_1c_45."Индикатор: Недолет" := FALSE;
   L_1c_45."Индикатор: Обрыв" := FALSE;
   L_1c_45."Индикатор: В норме" := FALSE;
   L_1c_45."Индикатор: HH активирована" := FALSE;
   L_1c_45."Индикатор: H активирована" := FALSE;
   L_1c_45."Индикатор: L активирована" := FALSE;
   L_1c_45."Индикатор: LL активирована" := FALSE;
   L_1c_45."Уставка: MAX" := 950.0;
   L_1c_45."Уставка: MIN" := 0.0;
   L_1c_45."Уставка: HH" := 80.0;
   L_1c_45."Уставка: H" := 70.0;
   L_1c_45."Уставка: L" := 15.0;
   L_1c_45."Уставка: LL" := 10.0;
   L_1c_45."Уставка: Перелёт" := 20.0;